// TIA Portal project "UploadAG314C_tia" (V15) (continued)
      STAT2038 : DInt;
      STAT2039 : DInt;
      STAT2040 : DInt;
      STAT2041 : DInt;
      STAT2042 : DInt;
      STAT2043 : Int;
      STAT2044 : Int := 100;
      STAT2045 : String[10];
      STAT2046 : DInt;
      STAT2047 : DInt;
      STAT2048 : DInt;
      STAT2049 : DInt;
      STAT2050 : DInt;
      STAT2051 : DInt;
      STAT2052 : DInt;
      STAT2053 : DInt;
      STAT2054 : DInt;
      STAT2055 : DInt;
      STAT2056 : DInt;
      STAT2057 : Int;
      STAT2058 : Int := 100;
      STAT2059 : String[10];
      STAT2060 : DInt;
      STAT2061 : DInt;
      STAT2062 : DInt;
      STAT2063 : DInt;
      STAT2064 : DInt;
      STAT2065 : DInt;
      STAT2066 : DInt;
      STAT2067 : DInt;
      STAT2068 : DInt;
      STAT2069 : DInt;
      STAT2070 : DInt;
      STAT2071 : Int;
      STAT2072 : Int := 100;
      STAT2073 : String[10];
      STAT2074 : DInt;
      STAT2075 : DInt;
      STAT2076 : DInt;
      STAT2077 : DInt;
      STAT2078 : DInt;
      STAT2079 : DInt;
      STAT2080 : DInt;
      STAT2081 : DInt;
      STAT2082 : DInt;
      STAT2083 : DInt;
      STAT2084 : DInt;
      STAT2085 : Int;
      STAT2086 : Int := 100;
      STAT2087 : String[10];
      STAT2088 : DInt;
      STAT2089 : DInt;
      STAT2090 : DInt;
      STAT2091 : DInt;
      STAT2092 : DInt;
      STAT2093 : DInt;
      STAT2094 : DInt;
      STAT2095 : DInt;
      STAT2096 : DInt;
      STAT2097 : DInt;
      STAT2098 : DInt;
      STAT2099 : Int;
      STAT2100 : Int := 100;
      STAT2101 : String[10];
      STAT2102 : DInt;
      STAT2103 : DInt;
      STAT2104 : DInt;
      STAT2105 : DInt;
      STAT2106 : DInt;
      STAT2107 : DInt;
      STAT2108 : DInt;
      STAT2109 : DInt;
      STAT2110 : DInt;
      STAT2111 : DInt;
      STAT2112 : DInt;
      STAT2113 : Int;
      STAT2114 : Int := 100;
      STAT2115 : String[10];
      STAT2116 : DInt;
      STAT2117 : DInt;
      STAT2118 : DInt;
      STAT2119 : DInt;
      STAT2120 : DInt;
      STAT2121 : DInt;
      STAT2122 : DInt;
      STAT2123 : DInt;
      STAT2124 : DInt;
      STAT2125 : DInt;
      STAT2126 : DInt;
      STAT2127 : Int;
      STAT2128 : Int := 100;
      STAT2129 : String[10];
      STAT2130 : DInt;
      STAT2131 : DInt;
      STAT2132 : DInt;
      STAT2133 : DInt;
      STAT2134 : DInt;
      STAT2135 : DInt;
      STAT2136 : DInt;
      STAT2137 : DInt;
      STAT2138 : DInt;
      STAT2139 : DInt;
      STAT2140 : DInt;
      STAT2141 : Int;
      STAT2142 : Int := 100;
      STAT2143 : String[10];
      STAT2144 : DInt;
      STAT2145 : DInt;
      STAT2146 : DInt;
      STAT2147 : DInt;
      STAT2148 : DInt;
      STAT2149 : DInt;
      STAT2150 : DInt;
      STAT2151 : DInt;
      STAT2152 : DInt;
      STAT2153 : DInt;
      STAT2154 : DInt;
      STAT2155 : Int;
      STAT2156 : Int := 100;
      STAT2157 : String[10];
      STAT2158 : DInt;
      STAT2159 : DInt;
      STAT2160 : DInt;
      STAT2161 : DInt;
      STAT2162 : DInt;
      STAT2163 : DInt;
      STAT2164 : DInt;
      STAT2165 : DInt;
      STAT2166 : DInt;
      STAT2167 : DInt;
      STAT2168 : DInt;
      STAT2169 : Int;
      STAT2170 : Int := 100;
      STAT2171 : String[10];
      STAT2172 : DInt;
      STAT2173 : DInt;
      STAT2174 : DInt;
      STAT2175 : DInt;
      STAT2176 : DInt;
      STAT2177 : DInt;
      STAT2178 : DInt;
      STAT2179 : DInt;
      STAT2180 : DInt;
      STAT2181 : DInt;
      STAT2182 : DInt;
      STAT2183 : Int;
      STAT2184 : Int := 100;
      STAT2185 : String[10];
      STAT2186 : DInt;
      STAT2187 : DInt;
      STAT2188 : DInt;
      STAT2189 : DInt;
      STAT2190 : DInt;
      STAT2191 : DInt;
      STAT2192 : DInt;
      STAT2193 : DInt;
      STAT2194 : DInt;
      STAT2195 : DInt;
      STAT2196 : DInt;
      STAT2197 : Int;
      STAT2198 : Int := 100;
      STAT2199 : String[10];
      STAT2200 : DInt;
      STAT2201 : DInt;
      STAT2202 : DInt;
      STAT2203 : DInt;
      STAT2204 : DInt;
      STAT2205 : DInt;
      STAT2206 : DInt;
      STAT2207 : DInt;
      STAT2208 : DInt;
      STAT2209 : DInt;
      STAT2210 : DInt;
      STAT2211 : Int;
      STAT2212 : Int := 100;
      STAT2213 : String[10];
      STAT2214 : DInt;
      STAT2215 : DInt;
      STAT2216 : DInt;
      STAT2217 : DInt;
      STAT2218 : DInt;
      STAT2219 : DInt;
      STAT2220 : DInt;
      STAT2221 : DInt;
      STAT2222 : DInt;
      STAT2223 : DInt;
      STAT2224 : DInt;
      STAT2225 : Int;
      STAT2226 : Int := 100;
      STAT2227 : String[10];
      STAT2228 : DInt;
      STAT2229 : DInt;
      STAT2230 : DInt;
      STAT2231 : DInt;
      STAT2232 : DInt;
      STAT2233 : DInt;
      STAT2234 : DInt;
      STAT2235 : DInt;
      STAT2236 : DInt;
      STAT2237 : DInt;
      STAT2238 : DInt;
      STAT2239 : Int;
      STAT2240 : Int := 100;
      STAT2241 : String[10];
      STAT2242 : DInt;
      STAT2243 : DInt;
      STAT2244 : DInt;
      STAT2245 : DInt;
      STAT2246 : DInt;
      STAT2247 : DInt;
      STAT2248 : DInt;
      STAT2249 : DInt;
      STAT2250 : DInt;
      STAT2251 : DInt;
      STAT2252 : DInt;
      STAT2253 : Int;
      STAT2254 : Int := 100;
      STAT2255 : String[10];
      STAT2256 : DInt;
      STAT2257 : DInt;
      STAT2258 : DInt;
      STAT2259 : DInt;
      STAT2260 : DInt;
      STAT2261 : DInt;
      STAT2262 : DInt;
      STAT2263 : DInt;
      STAT2264 : DInt;
      STAT2265 : DInt;
      STAT2266 : DInt;
      STAT2267 : Int;
      STAT2268 : Int := 100;
      STAT2269 : String[10];
      STAT2270 : DInt;
      STAT2271 : DInt;
      STAT2272 : DInt;
      STAT2273 : DInt;
      STAT2274 : DInt;
      STAT2275 : DInt;
      STAT2276 : DInt;
      STAT2277 : DInt;
      STAT2278 : DInt;
      STAT2279 : DInt;
      STAT2280 : DInt;
      STAT2281 : Int;
      STAT2282 : Int := 100;
      STAT2283 : String[10];
      STAT2284 : DInt;
      STAT2285 : DInt;
      STAT2286 : DInt;
      STAT2287 : DInt;
      STAT2288 : DInt;
      STAT2289 : DInt;
      STAT2290 : DInt;
      STAT2291 : DInt;
      STAT2292 : DInt;
      STAT2293 : DInt;
      STAT2294 : DInt;
      STAT2295 : Int;
      STAT2296 : Int := 100;
      STAT2297 : String[10];
      STAT2298 : DInt;
      STAT2299 : DInt;
      STAT2300 : DInt;
      STAT2301 : DInt;
      STAT2302 : DInt;
      STAT2303 : DInt;
      STAT2304 : DInt;
      STAT2305 : DInt;
      STAT2306 : DInt;
      STAT2307 : DInt;
      STAT2308 : DInt;
      STAT2309 : Int;
      STAT2310 : Int := 100;
      STAT2311 : String[10];
      STAT2312 : DInt;
      STAT2313 : DInt;
      STAT2314 : DInt;
      STAT2315 : DInt;
      STAT2316 : DInt;
      STAT2317 : DInt;
      STAT2318 : DInt;
      STAT2319 : DInt;
      STAT2320 : DInt;
      STAT2321 : DInt;
      STAT2322 : DInt;
      STAT2323 : Int;
      STAT2324 : Int := 100;
      STAT2325 : String[10];
      STAT2326 : DInt;
      STAT2327 : DInt;
      STAT2328 : DInt;
      STAT2329 : DInt;
      STAT2330 : DInt;
      STAT2331 : DInt;
      STAT2332 : DInt;
      STAT2333 : DInt;
      STAT2334 : DInt;
      STAT2335 : DInt;
      STAT2336 : DInt;
      STAT2337 : Int;
      STAT2338 : Int := 100;
      STAT2339 : String[10];
      STAT2340 : DInt;
      STAT2341 : DInt;
      STAT2342 : DInt;
      STAT2343 : DInt;
      STAT2344 : DInt;
      STAT2345 : DInt;
      STAT2346 : DInt;
      STAT2347 : DInt;
      STAT2348 : DInt;
      STAT2349 : DInt;
      STAT2350 : DInt;
      STAT2351 : Int;
      STAT2352 : Int := 100;
      STAT2353 : String[10];
      STAT2354 : DInt;
      STAT2355 : DInt;
      STAT2356 : DInt;
      STAT2357 : DInt;
      STAT2358 : DInt;
      STAT2359 : DInt;
      STAT2360 : DInt;
      STAT2361 : DInt;
      STAT2362 : DInt;
      STAT2363 : DInt;
      STAT2364 : DInt;
      STAT2365 : Int;
      STAT2366 : Int := 100;
      STAT2367 : String[10];
      STAT2368 : DInt;
      STAT2369 : DInt;
      STAT2370 : DInt;
      STAT2371 : DInt;
      STAT2372 : DInt;
      STAT2373 : DInt;
      STAT2374 : DInt;
      STAT2375 : DInt;
      STAT2376 : DInt;
      STAT2377 : DInt;
      STAT2378 : DInt;
      STAT2379 : Int;
      STAT2380 : Int := 100;
      STAT2381 : String[10];
      STAT2382 : DInt;
      STAT2383 : DInt;
      STAT2384 : DInt;
      STAT2385 : DInt;
      STAT2386 : DInt;
      STAT2387 : DInt;
      STAT2388 : DInt;
      STAT2389 : DInt;
      STAT2390 : DInt;
      STAT2391 : DInt;
      STAT2392 : DInt;
      STAT2393 : Int;
      STAT2394 : Int := 100;
      STAT2395 : String[10];
      STAT2396 : DInt;
      STAT2397 : DInt;
      STAT2398 : DInt;
      STAT2399 : DInt;
      STAT2400 : DInt;
      STAT2401 : DInt;
      STAT2402 : DInt;
      STAT2403 : DInt;
      STAT2404 : DInt;
      STAT2405 : DInt;
      STAT2406 : DInt;
      STAT2407 : Int;
      STAT2408 : Int := 100;
      STAT2409 : String[10];
      STAT2410 : DInt;
      STAT2411 : DInt;
      STAT2412 : DInt;
      STAT2413 : DInt;
      STAT2414 : DInt;
      STAT2415 : DInt;
      STAT2416 : DInt;
      STAT2417 : DInt;
      STAT2418 : DInt;
      STAT2419 : DInt;
      STAT2420 : DInt;
      STAT2421 : Int;
      STAT2422 : Int := 100;
      STAT2423 : String[10];
      STAT2424 : DInt;
      STAT2425 : DInt;
      STAT2426 : DInt;
      STAT2427 : DInt;
      STAT2428 : DInt;
      STAT2429 : DInt;
      STAT2430 : DInt;
      STAT2431 : DInt;
      STAT2432 : DInt;
      STAT2433 : DInt;
      STAT2434 : DInt;
      STAT2435 : Int;
      STAT2436 : Int := 100;
      STAT2437 : String[10];
      STAT2438 : DInt;
      STAT2439 : DInt;
      STAT2440 : DInt;
      STAT2441 : DInt;
      STAT2442 : DInt;
      STAT2443 : DInt;
      STAT2444 : DInt;
      STAT2445 : DInt;
      STAT2446 : DInt;
      STAT2447 : DInt;
      STAT2448 : DInt;
      STAT2449 : Int;
      STAT2450 : Int := 100;
      STAT2451 : String[10];
      STAT2452 : DInt;
      STAT2453 : DInt;
      STAT2454 : DInt;
      STAT2455 : DInt;
      STAT2456 : DInt;
      STAT2457 : DInt;
      STAT2458 : DInt;
      STAT2459 : DInt;
      STAT2460 : DInt;
      STAT2461 : DInt;
      STAT2462 : DInt;
      STAT2463 : Int;
      STAT2464 : Int := 100;
      STAT2465 : String[10];
      STAT2466 : DInt;
      STAT2467 : DInt;
      STAT2468 : DInt;
      STAT2469 : DInt;
      STAT2470 : DInt;
      STAT2471 : DInt;
      STAT2472 : DInt;
      STAT2473 : DInt;
      STAT2474 : DInt;
      STAT2475 : DInt;
      STAT2476 : DInt;
      STAT2477 : Int;
      STAT2478 : Int := 100;
      STAT2479 : String[10];
      STAT2480 : DInt;
      STAT2481 : DInt;
      STAT2482 : DInt;
      STAT2483 : DInt;
      STAT2484 : DInt;
      STAT2485 : DInt;
      STAT2486 : DInt;
      STAT2487 : DInt;
      STAT2488 : DInt;
      STAT2489 : DInt;
      STAT2490 : DInt;
      STAT2491 : Int;
      STAT2492 : Int := 100;
      STAT2493 : String[10];
      STAT2494 : DInt;
      STAT2495 : DInt;
      STAT2496 : DInt;
      STAT2497 : DInt;
      STAT2498 : DInt;
      STAT2499 : DInt;
      STAT2500 : DInt;
      STAT2501 : DInt;
      STAT2502 : DInt;
      STAT2503 : DInt;
      STAT2504 : DInt;
      STAT2505 : Int;
      STAT2506 : Int := 100;
      STAT2507 : String[10];
      STAT2508 : DInt;
      STAT2509 : DInt;
      STAT2510 : DInt;
      STAT2511 : DInt;
      STAT2512 : DInt;
      STAT2513 : DInt;
      STAT2514 : DInt;
      STAT2515 : DInt;
      STAT2516 : DInt;
      STAT2517 : DInt;
      STAT2518 : DInt;
      STAT2519 : Int;
      STAT2520 : Int := 100;
      STAT2521 : String[10];
      STAT2522 : DInt;
      STAT2523 : DInt;
      STAT2524 : DInt;
      STAT2525 : DInt;
      STAT2526 : DInt;
      STAT2527 : DInt;
      STAT2528 : DInt;
      STAT2529 : DInt;
      STAT2530 : DInt;
      STAT2531 : DInt;
      STAT2532 : DInt;
      STAT2533 : Int;
      STAT2534 : Int := 100;
      STAT2535 : String[10];
      STAT2536 : DInt;
      STAT2537 : DInt;
      STAT2538 : DInt;
      STAT2539 : DInt;
      STAT2540 : DInt;
      STAT2541 : DInt;
      STAT2542 : DInt;
      STAT2543 : DInt;
      STAT2544 : DInt;
      STAT2545 : DInt;
      STAT2546 : DInt;
      STAT2547 : Int;
      STAT2548 : Int := 100;
      STAT2549 : String[10];
      STAT2550 : DInt;
      STAT2551 : DInt;
      STAT2552 : DInt;
      STAT2553 : DInt;
      STAT2554 : DInt;
      STAT2555 : DInt;
      STAT2556 : DInt;
      STAT2557 : DInt;
      STAT2558 : DInt;
      STAT2559 : DInt;
      STAT2560 : DInt;
      STAT2561 : Int;
      STAT2562 : Int := 100;
      STAT2563 : String[10];
      STAT2564 : DInt;
      STAT2565 : DInt;
      STAT2566 : DInt;
      STAT2567 : DInt;
      STAT2568 : DInt;
      STAT2569 : DInt;
      STAT2570 : DInt;
      STAT2571 : DInt;
      STAT2572 : DInt;
      STAT2573 : DInt;
      STAT2574 : DInt;
      STAT2575 : Int;
      STAT2576 : Int := 100;
      STAT2577 : String[10];
      STAT2578 : DInt;
      STAT2579 : DInt;
      STAT2580 : DInt;
      STAT2581 : DInt;
      STAT2582 : DInt;
      STAT2583 : DInt;
      STAT2584 : DInt;
      STAT2585 : DInt;
      STAT2586 : DInt;
      STAT2587 : DInt;
      STAT2588 : DInt;
      STAT2589 : Int;
      STAT2590 : Int := 100;
      STAT2591 : String[10];
      STAT2592 : DInt;
      STAT2593 : DInt;
      STAT2594 : DInt;
      STAT2595 : DInt;
      STAT2596 : DInt;
      STAT2597 : DInt;
      STAT2598 : DInt;
      STAT2599 : DInt;
      STAT2600 : DInt;
      STAT2601 : DInt;
      STAT2602 : DInt;
      STAT2603 : Int;
      STAT2604 : Int := 100;
      STAT2605 : String[10];
      STAT2606 : DInt;
      STAT2607 : DInt;
      STAT2608 : DInt;
      STAT2609 : DInt;
      STAT2610 : DInt;
      STAT2611 : DInt;
      STAT2612 : DInt;
      STAT2613 : DInt;
      STAT2614 : DInt;
      STAT2615 : DInt;
      STAT2616 : DInt;
      STAT2617 : Int;
      STAT2618 : Int := 100;
      STAT2619 : String[10];
      STAT2620 : DInt;
      STAT2621 : DInt;
      STAT2622 : DInt;
      STAT2623 : DInt;
      STAT2624 : DInt;
      STAT2625 : DInt;
      STAT2626 : DInt;
      STAT2627 : DInt;
      STAT2628 : DInt;
      STAT2629 : DInt;
      STAT2630 : DInt;
      STAT2631 : Int;
      STAT2632 : Int := 100;
      STAT2633 : String[10];
      STAT2634 : DInt;
      STAT2635 : DInt;
      STAT2636 : DInt;
      STAT2637 : DInt;
      STAT2638 : DInt;
      STAT2639 : DInt;
      STAT2640 : DInt;
      STAT2641 : DInt;
      STAT2642 : DInt;
      STAT2643 : DInt;
      STAT2644 : DInt;
      STAT2645 : Int;
      STAT2646 : Int := 100;
      STAT2647 : String[10];
      STAT2648 : DInt;
      STAT2649 : DInt;
      STAT2650 : DInt;
      STAT2651 : DInt;
      STAT2652 : DInt;
      STAT2653 : DInt;
      STAT2654 : DInt;
      STAT2655 : DInt;
      STAT2656 : DInt;
      STAT2657 : DInt;
      STAT2658 : DInt;
      STAT2659 : Int;
      STAT2660 : Int := 100;
      STAT2661 : String[10];
      STAT2662 : DInt;
      STAT2663 : DInt;
      STAT2664 : DInt;
      STAT2665 : DInt;
      STAT2666 : DInt;
      STAT2667 : DInt;
      STAT2668 : DInt;
      STAT2669 : DInt;
      STAT2670 : DInt;
      STAT2671 : DInt;
      STAT2672 : DInt;
      STAT2673 : Int;
      STAT2674 : Int := 100;
      STAT2675 : String[10];
      STAT2676 : DInt;
      STAT2677 : DInt;
      STAT2678 : DInt;
      STAT2679 : DInt;
      STAT2680 : DInt;
      STAT2681 : DInt;
      STAT2682 : DInt;
      STAT2683 : DInt;
      STAT2684 : DInt;
      STAT2685 : DInt;
      STAT2686 : DInt;
      STAT2687 : Int;
      STAT2688 : Int := 100;
      STAT2689 : String[10];
      STAT2690 : DInt;
      STAT2691 : DInt;
      STAT2692 : DInt;
      STAT2693 : DInt;
      STAT2694 : DInt;
      STAT2695 : DInt;
      STAT2696 : DInt;
      STAT2697 : DInt;
      STAT2698 : DInt;
      STAT2699 : DInt;
      STAT2700 : DInt;
      STAT2701 : Int;
      STAT2702 : Int := 100;
      STAT2703 : String[10];
      STAT2704 : DInt;
      STAT2705 : DInt;
      STAT2706 : DInt;
      STAT2707 : DInt;
      STAT2708 : DInt;
      STAT2709 : DInt;
      STAT2710 : DInt;
      STAT2711 : DInt;
      STAT2712 : DInt;
      STAT2713 : DInt;
      STAT2714 : DInt;
      STAT2715 : Int;
      STAT2716 : Int := 100;
      STAT2717 : String[10];
      STAT2718 : DInt;
      STAT2719 : DInt;
      STAT2720 : DInt;
      STAT2721 : DInt;
      STAT2722 : DInt;
      STAT2723 : DInt;
      STAT2724 : DInt;
      STAT2725 : DInt;
      STAT2726 : DInt;
      STAT2727 : DInt;
      STAT2728 : DInt;
      STAT2729 : Int;
      STAT2730 : Int := 100;
      STAT2731 : String[10];
      STAT2732 : DInt;
      STAT2733 : DInt;
      STAT2734 : DInt;
      STAT2735 : DInt;
      STAT2736 : DInt;
      STAT2737 : DInt;
      STAT2738 : DInt;
      STAT2739 : DInt;
      STAT2740 : DInt;
      STAT2741 : DInt;
      STAT2742 : DInt;
      STAT2743 : Int;
      STAT2744 : Int := 100;
      STAT2745 : String[10];
      STAT2746 : DInt;
      STAT2747 : DInt;
      STAT2748 : DInt;
      STAT2749 : DInt;
      STAT2750 : DInt;
      STAT2751 : DInt;
      STAT2752 : DInt;
      STAT2753 : DInt;
      STAT2754 : DInt;
      STAT2755 : DInt;
      STAT2756 : DInt;
      STAT2757 : Int;
      STAT2758 : Int := 100;
      STAT2759 : String[10];
      STAT2760 : DInt;
      STAT2761 : DInt;
      STAT2762 : DInt;
      STAT2763 : DInt;
      STAT2764 : DInt;
      STAT2765 : DInt;
      STAT2766 : DInt;
      STAT2767 : DInt;
      STAT2768 : DInt;
      STAT2769 : DInt;
      STAT2770 : DInt;
      STAT2771 : Int;
      STAT2772 : Int := 100;
      STAT2773 : String[10];
      STAT2774 : DInt;
      STAT2775 : DInt;
      STAT2776 : DInt;
      STAT2777 : DInt;
      STAT2778 : DInt;
      STAT2779 : DInt;
      STAT2780 : DInt;
      STAT2781 : DInt;
      STAT2782 : DInt;
      STAT2783 : DInt;
      STAT2784 : DInt;
      STAT2785 : Int;
      STAT2786 : Int := 100;
      STAT2787 : String[10];
      STAT2788 : DInt;
      STAT2789 : DInt;
      STAT2790 : DInt;
      STAT2791 : DInt;
      STAT2792 : DInt;
      STAT2793 : DInt;
      STAT2794 : DInt;
      STAT2795 : DInt;
      STAT2796 : DInt;
      STAT2797 : DInt;
      STAT2798 : DInt;
      STAT2799 : Int;
      STAT2800 : Int := 100;
      STAT2801 : String[10];
      STAT2802 : DInt;
      STAT2803 : DInt;
      STAT2804 : DInt;
      STAT2805 : DInt;
      STAT2806 : DInt;
      STAT2807 : DInt;
      STAT2808 : DInt;
      STAT2809 : DInt;
      STAT2810 : DInt;
      STAT2811 : DInt;
      STAT2812 : DInt;
      STAT2813 : Int;
   END_VAR
BEGIN
END_DATA_BLOCK

DATA_BLOCK "Sampling_Data"   // DB18
{ S7_Optimized_Access := 'FALSE' }
VERSION : 0.1
   VAR
      Data_1 : Array[0..600] of Int;
      Data_2 : Array[0..600] of Int;
      Data_3 : Array[0..600] of Int;
      Data_4 : Array[0..600] of Int;
   END_VAR
BEGIN
END_DATA_BLOCK

DATA_BLOCK "Sampling_Control"   // DB21
{ S7_Optimized_Access := 'FALSE' }
VERSION : 0.1
   VAR
      startSave : Bool;
      trigerControl : Bool;
      dataSave : Bool;
      startLoging : Bool;
      trigerLogging : Bool;
      clearData : Bool;
      Sampling_time : S5Time := S5T#10ms;
      trigger_stop_log : Bool;
      stop_log_cmd : Bool;
      enable_poly_1 : Bool;
      enable_poly_2 : Bool;
      enable_poly_3 : Bool;
      enable_poly_4 : Bool;
      enable_iso_1 : Bool;
      enable_iso_2 : Bool;
      enable_iso_3 : Bool;
      enable_iso_4 : Bool;
   END_VAR
BEGIN
END_DATA_BLOCK

DATA_BLOCK "Sampling_Datalog"   // DB22
{ S7_Optimized_Access := 'FALSE' }
VERSION : 0.1
   VAR
      Datalog_poly_1 : Int;
      Datalog_poly_2 : Int;
      Datalog_poly_3 : Int;
      Datalog_poly_4 : Int;
      Datalog_iso_1 : Int;
      Datalog_iso_2 : Int;
      Datalog_iso_3 : Int;
      Datalog_iso_4 : Int;
      Count_datalog : Int;
   END_VAR
BEGIN
END_DATA_BLOCK

DATA_BLOCK "DB76"   // DB76
{ S7_Optimized_Access := 'FALSE' }
AUTHOR : JRW
VERSION : 0.1
   VAR
      STAT0 : Real;
      STAT1 : Real := 15.0;
      STAT2 : Real;
      STAT3 : Real;
      STAT4 : Real;
      STAT5 : Real;
      STAT6 : Real;
      STAT7 : Real;
      STAT8 : Real;
      STAT9 : Real;
      STAT10 : Real := 1.0;
      STAT11 : Real := 1.0;
      STAT12 : Real := 1.0;
      STAT13 : Real := 1.0;
      STAT14 : Real;
      STAT15 : Real;
      STAT16 : Real;
      STAT17 : Real;
      STAT18 : Real;
      STAT19 : Real;
      STAT20 : Real;
      STAT21 : Real := 12.0;
      STAT22 : Real := 10.0;
      STAT23 : Real := 80.0;
      STAT24 : Real;
      STAT25 : Real;
      STAT26 : Real;
      STAT27 : Int;
      STAT28 : Word;
      STAT29 : Word;
      STAT30 : Word;
      STAT31 : Word;
      STAT32 : Word;
      STAT33 : Bool;
      STAT34 : Bool;
      STAT35 : Bool;
      STAT36 : Bool;
      STAT37 : Bool := TRUE;
      STAT38 : Bool := TRUE;
      STAT39 : Bool := TRUE;
      STAT40 : Bool := TRUE;
      STAT41 : Bool := TRUE;
      STAT42 : Bool := TRUE;
      STAT43 : Bool;
      STAT44 : Bool;
      STAT45 : Bool := TRUE;
      STAT46 : Bool;
      STAT47 : Bool;
      STAT48 : Bool;
      STAT49 : Word;
      STAT50 : Word;
      STAT51 : Word;
      STAT52 : Int;
      STAT53 : Word;
      STAT54 : Word;
      STAT55 : Word := WORD#16#0015;
      STAT56 : Bool := TRUE;
      STAT57 : Int;
      STAT58 : Array[0..15] of Word;
      STAT59 : Array[0..4] of Word;
      STAT60 : Real := 0.88;
      STAT61 : Real := 1.025;
      STAT62 : Real := 1.094;
      STAT63 : Real := 1.093;
      STAT64 : Real := 0.934;
      STAT65 : Real := 1.075;
      STAT66 : Real := 1.0;
      STAT67 : Bool;
      STAT68 : Bool;
      STAT69 : Bool;
      STAT70 : Bool;
      STAT71 : Bool;
      STAT72 : Bool;
      STAT73 : Bool;
      STAT74 : Bool;
      STAT75 : Bool;
      STAT76 : Bool;
      STAT77 : Bool;
      STAT78 : Bool;
      STAT79 : Bool;
      STAT80 : Bool;
      STAT81 : Bool := TRUE;
      STAT82 : Bool;
      STAT83 : Bool;
      STAT84 : Bool;
      STAT85 : Bool;
      STAT86 : Bool;
      STAT87 : Bool;
      STAT88 : Bool;
      STAT89 : Bool;
      STAT90 : Bool;
      STAT91 : Bool;
      STAT92 : Int;
      STAT93 : Int := 50;
      STAT94 : Int := 5;
      STAT95 : Time := T#200MS;
      STAT96 : S5Time := S5T#1S;
      STAT97 : Date_And_Time;
      STAT98 : Bool;
      STAT99 : Bool;
      STAT100 : Real := 1.0;
      STAT101 : Real;
      STAT102 : Real;
      STAT103 : Bool;
      STAT104 : Int;
      STAT105 : Bool;
      STAT106 : Bool;
      STAT107 : Real;
      STAT108 : Real;
      STAT109 : Real;
      STAT110 : Real;
      STAT111 : Real;
      STAT112 : Real;
      STAT113 : Real;
      STAT114 : Real;
      STAT115 : Bool;
      STAT116 : Int;
      STAT117 : Word;
      STAT118 : Real;
      STAT119 : Real;
      STAT120 : Bool;
      STAT121 : Real;
      STAT122 : Word;
      STAT123 : Int;
      STAT124 : Word;
      STAT125 : Real;
      STAT126 : Word;
      STAT127 : Real;
      STAT128 : Bool;
      STAT129 : Bool;
      STAT130 : Bool;
      STAT131 : Bool;
      STAT132 : Int;
      STAT133 : String[16] := 'Entry';
      STAT134 : String[16] := 'Entry';
      STAT135 : String[16] := 'Entry';
      STAT136 : String[16] := 'Entry';
      STAT137 : Int;
      STAT138 : Int;
      STAT139 : Int;
      STAT140 : Int;
      STAT141 : Int;
      STAT142 : String[16] := 'Entry';
      STAT143 : Int;
      STAT144 : Int;
      STAT145 : Time := T#100MS;
      STAT146 : Time := T#5S;
      STAT147 : Time;
      STAT148 : Real := 1.6;
      STAT149 : Real := 40.0;
      STAT150 : Real := 2.0;
      STAT151 : Real := 37.5;
      STAT152 : Real := 31.3432;
      STAT153 : Real := 70.0;
      STAT154 : Real;
      STAT155 : Real;
      STAT156 : Real := 0.75;
      STAT157 : Real := 1.0;
      STAT158 : Real;
      STAT159 : Real;
      STAT160 : Bool;
   END_VAR
BEGIN
END_DATA_BLOCK

FUNCTION_BLOCK "FB1"   // FB1, LAD
{ S7_Optimized_Access := 'FALSE' }
VERSION : 0.1
   VAR_TEMP   // added for the SCL form of the ladder/FBD networks
      _w1 : Bool;
      _w2 : Bool;
      _s5time1 : S5Time;
   END_VAR
BEGIN

REGION Network 1 (STL)
         L     "Tag_4";
         DTR;
         L     "DB14".STAT21;
         DTR;
         *R;
         L     965.0;
         /R;
         L     9600.0;
         /R;
         RND;
         T     "DB12".STAT10;
         DTR;
         L     20.0;
         /R;
         T     "DB56".IN10;
END_REGION

REGION Network 2
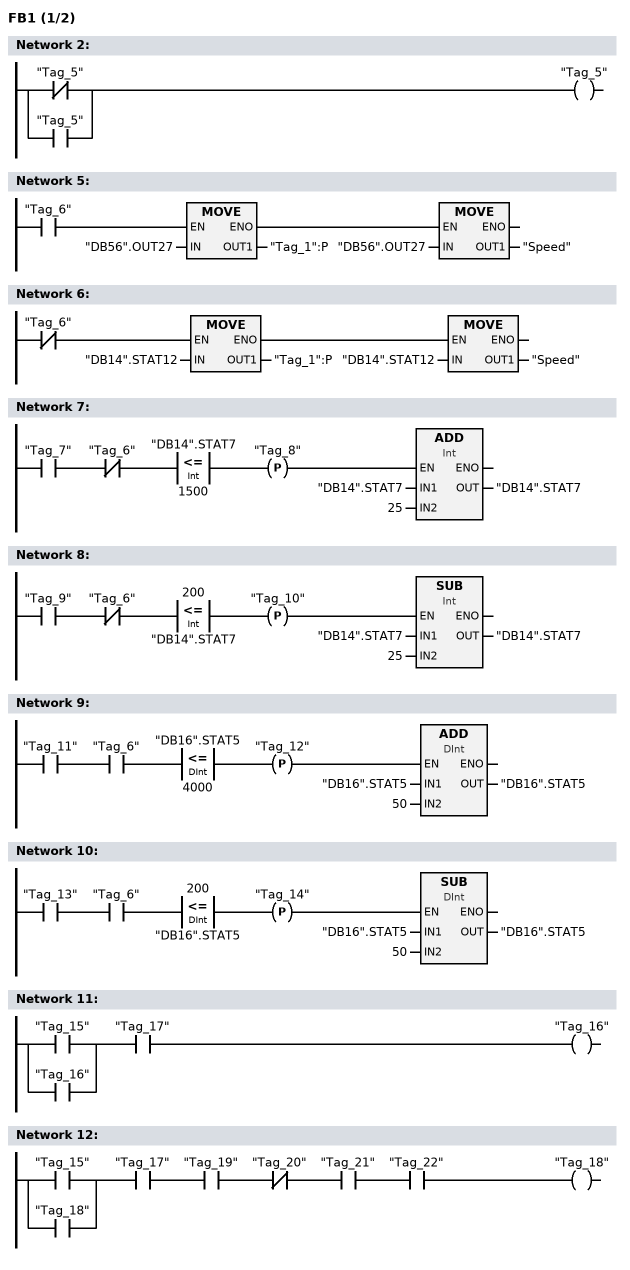
   RUNG wire#powerrail
      I_Contact( "Tag_5" )
      wire#w1
      Coil( "Tag_5" )
   END_RUNG
   RUNG wire#powerrail
      Contact( "Tag_5" )
   END_RUNG wire#w1
   // the same network as SCL:
   "Tag_5" := NOT "Tag_5" OR "Tag_5";
END_REGION

REGION Network 3 (STL)
         L     "DB16".STAT5;
         DTR;
         L     20.0;
         /R;
         T     "DB76".STAT151;
END_REGION

REGION Network 4 (STL)
         CALL  "FC51"
         ( IN0  := "DB14".STAT7,
           IN1  := 27648.0,
           IN2  := 0.0,
           IN3  := 1667.0,
           OUT4 := "DB14".STAT12
         );
         NOP   0;
END_REGION

REGION Network 5
   RUNG wire#powerrail
      Contact( "Tag_6" )
      { S7_GenerateENO := "TRUE" } Move(in := "DB56".OUT27, out1 => "Tag_1":P)
      { S7_GenerateENO := "TRUE" } Move(in := "DB56".OUT27, out1 => "Speed")
   END_RUNG
   // the same network as SCL:
   // ENO of a box is taken as its EN; it also drops when the box reports an error
   IF "Tag_6" THEN
       "Tag_1":P := "DB56".OUT27;
       "Speed" := "DB56".OUT27;
   END_IF;
END_REGION

REGION Network 6
   RUNG wire#powerrail
      I_Contact( "Tag_6" )
      { S7_GenerateENO := "TRUE" } Move(in := "DB14".STAT12, out1 => "Tag_1":P)
      { S7_GenerateENO := "TRUE" } Move(in := "DB14".STAT12, out1 => "Speed")
   END_RUNG
   // the same network as SCL:
   // ENO of a box is taken as its EN; it also drops when the box reports an error
   IF NOT "Tag_6" THEN
       "Tag_1":P := "DB14".STAT12;
       "Speed" := "DB14".STAT12;
   END_IF;
END_REGION

REGION Network 7
   RUNG wire#powerrail
      Contact( "Tag_7" )
      I_Contact( "Tag_6" )
      { S7_Templates := "SrcType := Int" } LE_Contact(in1 := "DB14".STAT7, in2 := 1500)
      P_Trig( "Tag_8" )
      { S7_Templates := "SrcType := Int"; S7_GenerateENO := "TRUE" } Add(in1 := "DB14".STAT7, in2 := 25, out => "DB14".STAT7)
   END_RUNG
   // the same network as SCL:
   #_w1 := "Tag_7" AND NOT "Tag_6" AND ("DB14".STAT7 <= 1500);
   #_w2 := #_w1 AND NOT "Tag_8";   // rising edge
   "Tag_8" := #_w1;
   IF #_w2 THEN "DB14".STAT7 := "DB14".STAT7 + 25; END_IF;
END_REGION

REGION Network 8
   RUNG wire#powerrail
      Contact( "Tag_9" )
      I_Contact( "Tag_6" )
      { S7_Templates := "SrcType := Int" } LE_Contact(in1 := 200, in2 := "DB14".STAT7)
      P_Trig( "Tag_10" )
      { S7_Templates := "SrcType := Int"; S7_GenerateENO := "TRUE" } Sub(in1 := "DB14".STAT7, in2 := 25, out => "DB14".STAT7)
   END_RUNG
   // the same network as SCL:
   #_w1 := "Tag_9" AND NOT "Tag_6" AND (200 <= "DB14".STAT7);
   #_w2 := #_w1 AND NOT "Tag_10";   // rising edge
   "Tag_10" := #_w1;
   IF #_w2 THEN "DB14".STAT7 := "DB14".STAT7 - 25; END_IF;
END_REGION

REGION Network 9
   RUNG wire#powerrail
      Contact( "Tag_11" )
      Contact( "Tag_6" )
      { S7_Templates := "SrcType := DInt" } LE_Contact(in1 := "DB16".STAT5, in2 := 4000)
      P_Trig( "Tag_12" )
      { S7_Templates := "SrcType := DInt"; S7_GenerateENO := "TRUE" } Add(in1 := "DB16".STAT5, in2 := 50, out => "DB16".STAT5)
   END_RUNG
   // the same network as SCL:
   #_w1 := "Tag_11" AND "Tag_6" AND ("DB16".STAT5 <= 4000);
   #_w2 := #_w1 AND NOT "Tag_12";   // rising edge
   "Tag_12" := #_w1;
   IF #_w2 THEN "DB16".STAT5 := "DB16".STAT5 + 50; END_IF;
END_REGION

REGION Network 10
   RUNG wire#powerrail
      Contact( "Tag_13" )
      Contact( "Tag_6" )
      { S7_Templates := "SrcType := DInt" } LE_Contact(in1 := 200, in2 := "DB16".STAT5)
      P_Trig( "Tag_14" )
      { S7_Templates := "SrcType := DInt"; S7_GenerateENO := "TRUE" } Sub(in1 := "DB16".STAT5, in2 := 50, out => "DB16".STAT5)
   END_RUNG
   // the same network as SCL:
   #_w1 := "Tag_13" AND "Tag_6" AND (200 <= "DB16".STAT5);
   #_w2 := #_w1 AND NOT "Tag_14";   // rising edge
   "Tag_14" := #_w1;
   IF #_w2 THEN "DB16".STAT5 := "DB16".STAT5 - 50; END_IF;
END_REGION

REGION Network 11
   RUNG wire#powerrail
      Contact( "Tag_15" )
      wire#w1
      Contact( "Tag_17" )
      Coil( "Tag_16" )
   END_RUNG
   RUNG wire#powerrail
      Contact( "Tag_16" )
   END_RUNG wire#w1
   // the same network as SCL:
   "Tag_16" := ("Tag_15" OR "Tag_16") AND "Tag_17";
END_REGION

REGION Network 12
   RUNG wire#powerrail
      Contact( "Tag_15" )
      wire#w1
      Contact( "Tag_17" )
      Contact( "Tag_19" )
      I_Contact( "Tag_20" )
      Contact( "Tag_21" )
      Contact( "Tag_22" )
      Coil( "Tag_18" )
   END_RUNG
   RUNG wire#powerrail
      Contact( "Tag_18" )
   END_RUNG wire#w1
   // the same network as SCL:
   "Tag_18" := ("Tag_15" OR "Tag_18") AND "Tag_17" AND "Tag_19" AND NOT "Tag_20" AND "Tag_21" AND "Tag_22";
END_REGION

REGION Network 13
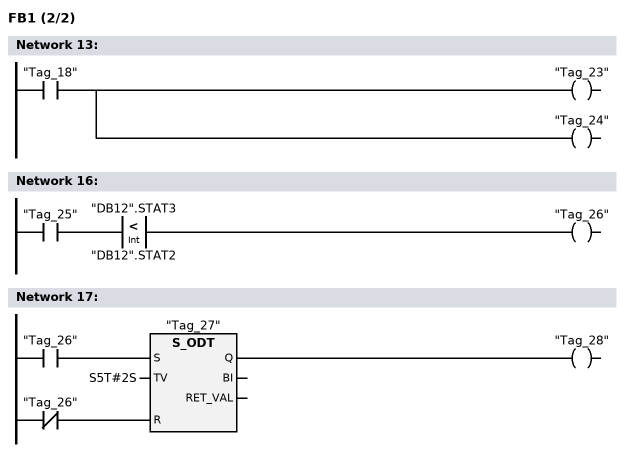
   RUNG wire#powerrail
      Contact( "Tag_18" )
      wire#w1
      Coil( "Tag_23" )
   END_RUNG
   RUNG wire#w1
      Coil( "Tag_24" )
   END_RUNG
   // the same network as SCL:
   "Tag_23" := "Tag_18";
   "Tag_24" := "Tag_18";
END_REGION

REGION Network 14 (STL)
         CALL  "FC52"
         ( IN0  := "Tag_2":P,
           IN1  := 900.0,
           IN2  := 0.0,
           OUT3 := "DB13".STAT7
         );
END_REGION

REGION Network 15 (STL)
         L     "Tag_3":P;
         T     "DB12".STAT3;
END_REGION

REGION Network 16
   RUNG wire#powerrail
      Contact( "Tag_25" )
      { S7_Templates := "SrcType := Int" } LT_Contact(in1 := "DB12".STAT3, in2 := "DB12".STAT2)
      Coil( "Tag_26" )
   END_RUNG
   // the same network as SCL:
   "Tag_26" := "Tag_25" AND ("DB12".STAT3 < "DB12".STAT2);
END_REGION

REGION Network 17
   RUNG wire#powerrail
      Contact( "Tag_26" )
      S_ODT(T_NO := "Tag_27", TV := S5T#2S, R := wire#w1, BI =>, RET_VAL =>)
      Coil( "Tag_28" )
   END_RUNG
   RUNG wire#powerrail
      I_Contact( "Tag_26" )
   END_RUNG wire#w1
   // the same network as SCL:
   #_s5time1 := S_ODT(T_NO := "Tag_27", TV := S5T#2S, S := "Tag_26", R := NOT "Tag_26", Q => #_w1);
   "Tag_28" := #_w1;
END_REGION
END_FUNCTION_BLOCK

FUNCTION "FC51" : Void   // FC51, STL
{ S7_Optimized_Access := 'FALSE' }
VERSION : 0.0
   VAR_INPUT
      IN0 : Int;
      IN1 : Real;
      IN2 : Real;
      IN3 : Real;
   END_VAR
   VAR_OUTPUT
      OUT4 : Int;
   END_VAR
   VAR_TEMP
      TEMP5 : Real;
      TEMP6 : Real;
   END_VAR
BEGIN

REGION Network 1
         L     #IN0;
         ITD;
         DTR;
         T     #TEMP5;
END_REGION

REGION Network 2
         L     #IN1;
         L     #IN2;
         -R;
         T     #TEMP6;
END_REGION

REGION Network 3
         L     #TEMP5;
         L     #IN3;
         /R;
         L     #TEMP6;
         *R;
         L     #IN2;
         +R;
         TRUNC;
         T     "Tag_29";
         L     "Tag_30";
         T     #OUT4;
END_REGION
END_FUNCTION

FUNCTION "FC52" : Void   // FC52, STL
{ S7_Optimized_Access := 'FALSE' }
VERSION : 0.0
   VAR_INPUT
      IN0 : Int;
      IN1 : Real;
      IN2 : Real;
   END_VAR
   VAR_OUTPUT
      OUT3 : Real;
   END_VAR
   VAR_TEMP
      TEMP4 : Real;
      TEMP5 : Real;
      TEMP6 : Real;
   END_VAR
BEGIN

REGION Network 1
         L     #IN0;
         ITD;
         DTR;
         T     #TEMP4;
END_REGION

REGION Network 2
         L     #TEMP4;
         L     65.5;
         -R;
         T     #TEMP5;
END_REGION

REGION Network 3
         L     #IN1;
         L     #IN2;
         -R;
         T     #TEMP6;
END_REGION

REGION Network 4
         L     #TEMP5;
         L     2764.8;
         /R;
         L     #TEMP6;
         *R;
         L     #IN2;
         +R;
         TRUNC;
         L     2;
         <=I;
         JC    M001;
         TAK;
         JU    M002;
   M001: L     0;
         T     #OUT3;
   M002: T     #OUT3;
END_REGION
END_FUNCTION

FUNCTION "Sampling_Execution" : Void   // FC353, LAD
TITLE = Sampling Execution
{ S7_Optimized_Access := 'FALSE' }
VERSION : 0.1
   VAR_TEMP   // added for the SCL form of the ladder/FBD networks
      _w1 : Bool;
      _s5time1 : S5Time;
      _w2 : Bool;
      _w3 : Bool;
      _w4 : Bool;
      _w5 : Bool;
      _w6 : Bool;
      _s5time2 : S5Time;
   END_VAR
BEGIN

REGION Network 1: Pressure Save data for sampling
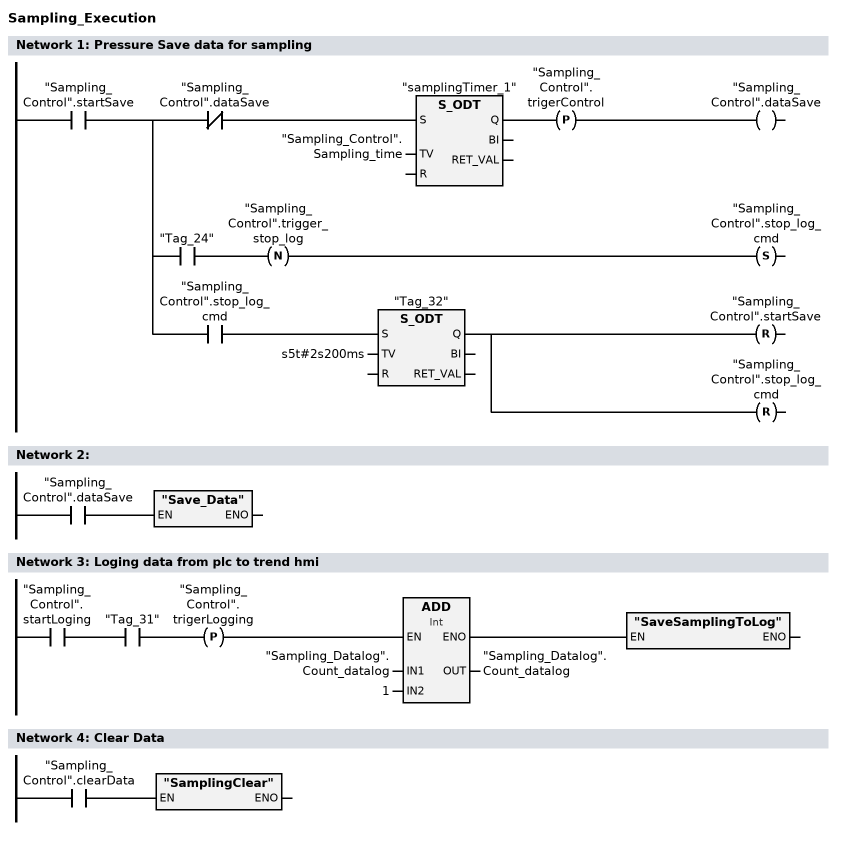
   RUNG wire#powerrail
      Contact( "Sampling_Control".startSave )
      wire#w1
      I_Contact( "Sampling_Control".dataSave )
      S_ODT(T_NO := "samplingTimer_1", TV := "Sampling_Control".Sampling_time, R :=, BI =>, RET_VAL =>)
      P_Trig( "Sampling_Control".trigerControl )
      Coil( "Sampling_Control".dataSave )
   END_RUNG
   RUNG wire#w1
      Contact( "Tag_24" )
      N_Trig( "Sampling_Control".trigger_stop_log )
      S_Coil( "Sampling_Control".stop_log_cmd )
   END_RUNG
   RUNG wire#w1
      Contact( "Sampling_Control".stop_log_cmd )
      S_ODT(T_NO := "Tag_32", TV := s5t#2s200ms, R :=, BI =>, RET_VAL =>)
      wire#w2
      R_Coil( "Sampling_Control".startSave )
   END_RUNG
   RUNG wire#w2
      R_Coil( "Sampling_Control".stop_log_cmd )
   END_RUNG
   // the same network as SCL:
   #_w2 := "Sampling_Control".startSave;
   #_s5time1 := S_ODT(T_NO := "samplingTimer_1",
                      S := "Sampling_Control".startSave AND NOT "Sampling_Control".dataSave,
                      TV := "Sampling_Control".Sampling_time,
                      Q => #_w1);
   #_w3 := #_w1 AND NOT "Sampling_Control".trigerControl;   // rising edge
   "Sampling_Control".trigerControl := #_w1;
   "Sampling_Control".dataSave := #_w3;
   #_w4 := #_w2 AND "Tag_24";
   #_w5 := NOT #_w4 AND "Sampling_Control".trigger_stop_log;   // falling edge
   "Sampling_Control".trigger_stop_log := #_w4;
   IF #_w5 THEN "Sampling_Control".stop_log_cmd := TRUE; END_IF;
   #_s5time2 := S_ODT(T_NO := "Tag_32",
                      S := #_w2 AND "Sampling_Control".stop_log_cmd,
                      TV := s5t#2s200ms,
                      Q => #_w6);
   IF #_w6 THEN
       "Sampling_Control".startSave := FALSE;
       "Sampling_Control".stop_log_cmd := FALSE;
   END_IF;
END_REGION

REGION Network 2
   RUNG wire#powerrail
      Contact( "Sampling_Control".dataSave )
      "Save_Data"()
   END_RUNG
   // the same network as SCL:
   IF "Sampling_Control".dataSave THEN "Save_Data"(); END_IF;
END_REGION

REGION Network 3: Loging data from plc to trend hmi
   RUNG wire#powerrail
      Contact( "Sampling_Control".startLoging )
      Contact( "Tag_31" )
      P_Trig( "Sampling_Control".trigerLogging )
      { S7_Templates := "SrcType := Int"; S7_GenerateENO := "TRUE" } Add(in1 := "Sampling_Datalog".Count_datalog, in2 := 1, out => "Sampling_Datalog".Count_datalog)
      "SaveSamplingToLog"()
   END_RUNG
   // the same network as SCL:
   // ENO of a box is taken as its EN; it also drops when the box reports an error
   #_w1 := "Sampling_Control".startLoging AND "Tag_31";
   #_w2 := #_w1 AND NOT "Sampling_Control".trigerLogging;   // rising edge
   "Sampling_Control".trigerLogging := #_w1;
   IF #_w2 THEN
       "Sampling_Datalog".Count_datalog := "Sampling_Datalog".Count_datalog + 1;
       "SaveSamplingToLog"();
   END_IF;
END_REGION

REGION Network 4: Clear Data
   RUNG wire#powerrail
      Contact( "Sampling_Control".clearData )
      "SamplingClear"()
   END_RUNG
   // the same network as SCL:
   IF "Sampling_Control".clearData THEN "SamplingClear"(); END_IF;
END_REGION
END_FUNCTION

FUNCTION "SaveSamplingToLog" : Void   // FC354, SCL
TITLE = save data dari sampling ke log
{ S7_Optimized_Access := 'FALSE' }
VERSION : 0.1
   VAR_TEMP
      x : Int;
   END_VAR
BEGIN

   IF "Sampling_Control".startLoging = TRUE THEN
       #x := 600 - "Sampling_Datalog".Count_datalog;
       //Pressure
       "Sampling_Datalog".Datalog_poly_1:= "Sampling_Data".Data_1[#x];
       //Flowrate
       "Sampling_Datalog".Datalog_poly_2 :="Sampling_Data".Data_2[#x];
       //Temperature
       "Sampling_Datalog".Datalog_poly_3 :="Sampling_Data".Data_3[#x];
       //speed
       "Sampling_Datalog".Datalog_poly_4 := "Sampling_Data".Data_4[#x];

       IF "Sampling_Datalog".Count_datalog >= 600 THEN

           "Sampling_Control".startLoging := FALSE;

       END_IF;
   END_IF;
END_FUNCTION

FUNCTION "SamplingClear" : Void   // FC355, SCL
TITLE = untuk clear sampling data
{ S7_Optimized_Access := 'FALSE' }
VERSION : 0.1
   VAR_TEMP
      i : Int;
   END_VAR
BEGIN
   FOR #i := 0 TO 600 DO
       "Sampling_Data".Data_1[#i] := 0;
       "Sampling_Data".Data_2[#i] := 0;
       "Sampling_Data".Data_3[#i] := 0;
       "Sampling_Data".Data_4[#i] := 0;

   END_FOR;
   "Sampling_Datalog".Datalog_poly_1 := 0;
   "Sampling_Datalog".Datalog_poly_2 := 0;
   "Sampling_Datalog".Datalog_poly_3 := 0;
   "Sampling_Datalog".Datalog_poly_4 := 0;


   "Sampling_Datalog".Count_datalog := 0;
   "Sampling_Control".clearData := FALSE;
END_FUNCTION

FUNCTION "Save_Data" : Void   // FC356, SCL
{ S7_Optimized_Access := 'FALSE' }
VERSION : 0.1
   VAR_TEMP
      i : Int;
   END_VAR
BEGIN
   REGION cntrl save
           FOR #i := (600 - 1) TO 0 BY -1 DO
               // Data 1 = Pressure
               "Sampling_Data".Data_1[#i + 1] := "Sampling_Data".Data_1[#i];
               "Sampling_Data".Data_2[#i + 1] := "Sampling_Data".Data_2[#i];
               "Sampling_Data".Data_3[#i + 1] := "Sampling_Data".Data_3[#i];
               "Sampling_Data".Data_4[#i + 1] := "Sampling_Data".Data_4[#i];

           END_FOR;


           REGION save data 1
               // Data 1 = Pressure
               IF "Sampling_Control".enable_poly_1 = TRUE THEN
                   "Sampling_Data".Data_1[0] := DINT_TO_INT(%DB12.DBD32);
               ELSE
                   "Sampling_Data".Data_1[0] := 0;
               END_IF;

             END_REGION
           REGION save data 2
               // Data 2 = Flowrate
               IF "Sampling_Control".enable_poly_2 = TRUE THEN
                   "Sampling_Data".Data_2[0] := DINT_TO_INT(%DB13.DBD28);
               ELSE
                   "Sampling_Data".Data_2[0] := 0;
               END_IF;

              END_REGION
           REGION save data 3
               // Data 3 = Temperature
               IF "Sampling_Control".enable_poly_3 = TRUE THEN
                   "Sampling_Data".Data_3[0] := %DB12.DBW6;
               ELSE
                   "Sampling_Data".Data_3[0] := 0;
               END_IF;
              END_REGION
           REGION save data 4
               // Data 4 = Speed
               IF "Sampling_Control".enable_poly_4 = TRUE THEN
                   "Sampling_Data".Data_4[0] := "Speed";
               ELSE
                   "Sampling_Data".Data_4[0] := 0;
               END_IF;
           END_REGION
     END_REGION
END_FUNCTION

ORGANIZATION_BLOCK "OB1"   // OB1, STL
{ S7_Optimized_Access := 'FALSE' }
VERSION : 0.1
   VAR_TEMP
      TEMP0 : Byte;
      TEMP1 : Byte;
      TEMP2 : Byte;
      TEMP3 : Byte;
      TEMP4 : Byte;
      TEMP5 : Byte;
      TEMP6 : Int;
      TEMP7 : Int;
      TEMP8 : Int;
      TEMP9 : Date_And_Time;
   END_VAR
BEGIN

REGION Network 1
         UC    "FB1";
END_REGION

REGION Network 2
         CALL  "Sampling_Execution";
END_REGION
END_ORGANIZATION_BLOCK

ORGANIZATION_BLOCK "OB35"   // OB35, STL
{ S7_Optimized_Access := 'FALSE' }
VERSION : 0.1
   VAR_TEMP
      TEMP0 : Byte;
      TEMP1 : Byte;
      TEMP2 : Byte;
      TEMP3 : Byte;
      TEMP4 : Byte;
      TEMP5 : Byte;
      TEMP6 : Word;
      TEMP7 : Int;
      TEMP8 : Int;
      TEMP9 : Date_And_Time;
   END_VAR
BEGIN

REGION Network 1
         CALL  FREQUENC_300C , "DB30"
         ( LADDR    := ,
           CHANNEL  := 0,
           SW_GATE  := "Tag_24",
           MAN_DO   := ,
           SET_DO   := ,
           JOB_REQ  := ,
           JOB_ID   := ,
           JOB_VAL  := ,
           STS_GATE := ,
           STS_STRT := ,
           STS_DO   := ,
           STS_C_DN := ,
           STS_C_UP := ,
           MEAS_VAL := "Tag_4",
           COUNTVAL := ,
           JOB_DONE := ,
           JOB_ERR  := ,
           JOB_STAT :=
         );
END_REGION

REGION Network 2
         AN    "Tag_24";
         =     %L20.0;
         BLD   103;
         A     "Tag_5";
         =     %L20.4;
         BLD   103;
         CALL  "CONT_C_LF", "DB56"
         ( IN0   := %L20.0,
           IN1   := ,
           IN2   := ,
           IN3   := FALSE,
           IN4   := %L20.4,
           IN5   := FALSE,
           IN6   := FALSE,
           IN7   := FALSE,
           IN8   := T#10MS,
           IN9   := "DB76".STAT151,
           IN10  := ,
           IN11  := ,
           IN12  := ,
           IN13  := "DB76".STAT148,
           IN14  := "DB76".STAT145,
           IN15  := T#1S,
           IN16  := T#200MS,
           IN17  := ,
           IN18  := ,
           IN19  := ,
           IN20  := ,
           IN21  := ,
           IN22  := ,
           IN23  := ,
           IN24  := ,
           IN25  := ,
           OUT26 := ,
           OUT27 := ,
           OUT28 := ,
           OUT29 := ,
           OUT30 := ,
           OUT31 := ,
           OUT32 := ,
           OUT33 := ,
           OUT34 :=
         );
         NOP   0;
END_REGION
END_ORGANIZATION_BLOCK

ORGANIZATION_BLOCK "OB80"   // OB80, LAD
{ S7_Optimized_Access := 'FALSE' }
VERSION : 0.1
   VAR_TEMP
      TEMP0 : Byte;
      TEMP1 : Byte;
      TEMP2 : Byte;
      TEMP3 : Byte;
      TEMP4 : Byte;
      TEMP5 : Byte;
      TEMP6 : Word;
      TEMP7 : Byte;
      TEMP8 : Byte;
      TEMP9 : Byte;
      TEMP10 : Byte;
      TEMP11 : Date_And_Time;
   END_VAR
BEGIN
END_ORGANIZATION_BLOCK

ORGANIZATION_BLOCK "OB82"   // OB82, LAD
{ S7_Optimized_Access := 'FALSE' }
VERSION : 0.1
   VAR_TEMP
      TEMP0 : Byte;
      TEMP1 : Byte;
      TEMP2 : Byte;
      TEMP3 : Byte;
      TEMP4 : Byte;
      TEMP5 : Byte;
      TEMP6 : Word;
      TEMP7 : Bool;
      TEMP8 : Bool;
      TEMP9 : Bool;
      TEMP10 : Bool;
      TEMP11 : Bool;
      TEMP12 : Bool;
      TEMP13 : Bool;
      TEMP14 : Bool;
      TEMP15 : Byte;
      TEMP16 : Bool;
      TEMP17 : Bool;
      TEMP18 : Bool;
      TEMP19 : Bool;
      TEMP20 : Bool;
      TEMP21 : Bool;
      TEMP22 : Bool;
      TEMP23 : Bool;
      TEMP24 : Bool;
      TEMP25 : Bool;
      TEMP26 : Bool;
      TEMP27 : Bool;
      TEMP28 : Bool;
      TEMP29 : Bool;
      TEMP30 : Bool;
      TEMP31 : Bool;
      TEMP32 : Date_And_Time;
   END_VAR
BEGIN
END_ORGANIZATION_BLOCK

ORGANIZATION_BLOCK "OB121"   // OB121, LAD
{ S7_Optimized_Access := 'FALSE' }
VERSION : 0.1
   VAR_TEMP
      TEMP0 : Byte;
      TEMP1 : Byte;
      TEMP2 : Byte;
      TEMP3 : Byte;
      TEMP4 : Byte;
      TEMP5 : Byte;
      TEMP6 : Word;
      TEMP7 : Word;
      TEMP8 : Word;
      TEMP9 : Date_And_Time;
   END_VAR
BEGIN
END_ORGANIZATION_BLOCK

ORGANIZATION_BLOCK "OB122"   // OB122, LAD
{ S7_Optimized_Access := 'FALSE' }
VERSION : 0.1
   VAR_TEMP
      TEMP0 : Byte;
      TEMP1 : Byte;
      TEMP2 : Byte;
      TEMP3 : Byte;
      TEMP4 : Byte;
      TEMP5 : Byte;
      TEMP6 : Word;
      TEMP7 : Word;
      TEMP8 : Word;
      TEMP9 : Date_And_Time;
   END_VAR
BEGIN
END_ORGANIZATION_BLOCK

(* ===== HMI "HMI_RT_2" =====
system functions are stored by id; their names below are inferred from use
connection "SPS_1": IF1 B, SIMATIC S7 300/400 MPI

HMI tags "Default tag table"
   "NavUserChange" : Int, internal
   "NavScreenChange" : Int, internal
   "Alarm_Filter_Tag" : Int, internal
   "tes_1" : Bool, internal
   "tes_2" : Bool, internal
   "tes_3" : Bool, internal
   "Date_1" : DateTime, internal
   "Date" : DateTime, internal
   "Time" : DateTime, internal
   "HMI_Tag_1" : Int, internal
   "HMI_Tag_1(1)" : Int, internal
   "tes_Time_1" : DateTime, internal
   "tes_Time_2" : DateTime, internal
   "tes_Time_3" : DateTime, internal
   "Shot" : Bool AT %DB205.DBX122.1, 1 s
   "Meter" : Bool AT %DB30.DBX112.7, 1 s
   "Cycle" : Bool AT %DB205.DBX122.0, 1 s
   "Bar_1" : Bool AT %DB205.DBX122.2, 1 s
   "safely_remove_usb" : Bool, internal
   "CopyfromSD" : Bool, internal
   "CopyfromUSB" : Bool, internal
   "Anim_OpenLOgs" : Bool, internal

HMI tags "Sampling_Trend"
   "saveDataControl" : Bool AT %DB21.DBX0.0, 1 s
   "loggingDataControl" : Bool AT %DB21.DBX0.3, 1 s
   "count" : Int AT %DB22.DBW16, 100 ms
      on ChangeValue: "StartStopLogging"()
   "pressure_poly" : Int AT %DB22.DBW0, 100 ms
      on ChangeValue: function_abcfba0d("temperature_poly"); function_abcfba0d("temperature_iso")
   "flowrate_poly" : Int AT %DB22.DBW2, 100 ms
      on ChangeValue: function_abcfba0d("speed_poly")
   "temperature_poly" : Int AT %DB22.DBW4, 100 ms
   "cleardata" : Bool AT %DB21.DBX0.5, 1 s
   "savetrend" : Int, internal
   "loadtrend" : Int, internal
   "pressure_iso" : Int AT %DB22.DBW8, 100 ms
   "flowrate_iso" : Int AT %DB22.DBW10, 100 ms
   "temperature_iso" : Int AT %DB22.DBW12, 100 ms
   "fileChossen" : WString[200], internal
   "archive_path" : WString[200], internal
   "current_dir" : WString[200], internal
   "count_res" : Int, internal
   "flowrate_iso_res" : Int, internal
   "flowrate_poly_res" : Int, internal
   "pressure_poly_res" : Int, internal
   "pressure_iso_res" : Int, internal
   "stat_fileChosen" : Int, internal
   "restore_time" : DateTime, internal
   "Trend_startingTime" : DateTime, internal
   "Trend_endTime" : DateTime, internal
   "Trend_index" : Int, internal
   "trend_index2" : Int, internal
   "Sampling_Time" : S5Time AT %DB21.DBW2, 1 s
   "Sampling_Alarm" : Int, internal
   "temperature_poly_res" : Int, internal
   "temperature_iso_res" : Int, internal
   "PrintScreenButton" : Bool, internal
   "speed_poly" : Int AT %DB22.DBW6, 1 s
   "speed_poly_res" : Int, internal
   "speed_iso" : Int AT %DB22.DBW14, 1 s
   "speed_iso_res" : Int, internal
   "enable_poly_1" : Bool AT %DB21.DBX4.2, 1 s
   "enable_poly_2" : Bool AT %DB21.DBX4.3, 1 s
   "enable_poly_3" : Bool AT %DB21.DBX4.4, 1 s
   "enable_poly_4" : Bool AT %DB21.DBX4.5, 1 s
   "enable_iso_1" : Bool AT %DB21.DBX4.6, 1 s
   "enable_iso_2" : Bool AT %DB21.DBX4.7, 1 s
   "enable_iso_3" : Bool AT %DB21.DBX5.0, 1 s
   "enable_iso_4" : Bool AT %DB21.DBX5.1, 1 s

HMI tags "LHmiView_FileBrowser"
   "File_1" : WString[255], internal
   "File_10" : WString[255], internal
   "File_2" : WString[255], internal
   "File_3" : WString[255], internal
   "File_4" : WString[255], internal
   "File_5" : WString[255], internal
   "File_6" : WString[255], internal
   "File_7" : WString[255], internal
   "File_8" : WString[255], internal
   "File_9" : WString[255], internal
   "Folder" : WString[255], internal
   "isFolder_1" : WString[10], internal
   "isFolder_2" : WString[10], internal
   "isFolder_3" : WString[10], internal
   "isFolder_4" : WString[10], internal
   "isFolder_5" : WString[10], internal
   "isFolder_6" : WString[10], internal
   "isFolder_7" : WString[10], internal
   "isFolder_8" : WString[10], internal
   "isFolder_9" : WString[10], internal
   "isFolder_10" : WString[10], internal
   "NextPossible" : Bool, internal
   "index" : Int, internal
   "fileChosen" : Int, internal
   "NewFolder" : WString[255], internal
   "NewName" : WString[255], internal
   "bufferFile" : WString[255], internal
   "bufferFolder" : WString[255], internal
   "bufferIsFolder" : Bool, internal
   "bufferCopyCut" : Bool, internal
   "pdfPath" : WString[80], internal
   "htmlPath" : WString[80], internal
   "FEStatus" : WString[150], internal
   "FEsearchString" : WString[80], internal
   "Search" : Bool, internal
   "FEsearchFolder" : WString[80], internal
   "stateBackground" : Bool, internal

